(* Logix 5000 project; controller PLC_MCC1300_75F1 vendor 1 type 14 code 166 rev 32.11; software revision 32.04; part 75 of 83 *)
(* tags used below, declared in another part *)
   AUX_tBufferPlate_NULL : UDT_BufferPlate;
   AUX_tHMI_Lite_NULL : UDT_HMI_LITE;
   CONST_rgdDestMask : DINT[32];   // Destination Mask
   CONST_tPlant : UDT_PLANT_CONSTANTS;
   GP_OB_InitializeMain : GP_OB_Initialize;
   GP_PosWindow : GP_PosWindow;
   GP_RampManagement : GP_RampManagement;
   GP_RampSpace : GP_RampSpace;
   M30xTrimDeck : MAC_TrimmingDeck[5];
   M30xTrimDeck_HMR : MAC_TrimmingDeck_HMR[5];
   M30xTrimDeck_HMW : MAC_TrimmingDeck_HMW[5];
   M30xTrimWheel : MAC_TrimmingWheels[5];
   M30xTrimWheel_HMW : MAC_TrimmingWheels_HMW[5];
   M311_Data : UDT_Convoy_SL;
   M311A_Data : UDT_Convoy_SL;
   Sbr_IN_dCapIndex : DINT;
   Sbr_IN_dConveyor : DINT;
   Sbr_IN_DestinationCullet : DINT;
   Sbr_IN_DestinationID : DINT;
   Sbr_IN_dIndexHead : DINT;
   Sbr_IN_dMaskAllowed : DINT;
   Sbr_IN_Position : DINT;
   Sbr_IN_PosStart : DINT;
   Sbr_IN_PosStop : DINT;
   Sbr_IN_ReasonID : DINT;
   Sbr_IN_xHeadPos : BOOL;
   Sbr_IN_xSendAllCullet : BOOL;
   Sbr_INO_DestinationLite : DINT;
   Sbr_INO_tConvoy_SL : UDT_Convoy_SL;
   Sbr_OUT_dIndexTail : DINT;
   Sbr_OUT_ReqRot_CCW : BOOL;
   Sbr_OUT_ReqRot_CW : BOOL;
   TMP_d : DINT;
   TMP_d2 : DINT;
   TMP_dAccSpace : DINT;
   TMP_dActualSpeed : DINT;
   TMP_dBufferSize : DINT;
   TMP_dCap : DINT;
   TMP_dCapNextConvoy : DINT;
   TMP_dConveyorLength : DINT;
   TMP_dConvoySearchMax : DINT;
   TMP_dCountDest : DINT;
   TMP_dCulletMask : DINT;
   TMP_dDecSpace : DINT;
   TMP_dHeadMax : DINT;
   TMP_dHeadPosition_mm : DINT;
   TMP_dIndex : DINT;
   TMP_dIndex2 : DINT;
   TMP_dIndex3 : DINT;
   TMP_dIndex4 : DINT;
   TMP_dIndexCap : DINT;
   TMP_dIndexCapConv : DINT;
   TMP_dIndexConv : DINT;
   TMP_dIndexMotor : DINT;
   TMP_dIndexNext : DINT;
   TMP_dIndexPlate : DINT;
   TMP_dLastConv : DINT;
   TMP_dLastConvTail : DINT;
   TMP_dLineSize : DINT;
   TMP_dLite : DINT;
   TMP_dLiteInv : DINT;
   TMP_dManualTargetPos : DINT;
   TMP_dMask : DINT;
   TMP_dMaxCap : DINT;
   TMP_dMaxLite : DINT;
   TMP_dMinTail : DINT;
   TMP_dNextCap : DINT;
   TMP_dPointerCap : DINT;
   TMP_dPos_cmm : DINT;
   TMP_dPosHead_cmm : DINT;
   TMP_dPosTail_cmm : DINT;
   TMP_dRampMotor : DINT;
   TMP_dStepAdvMotor : DINT;
   TMP_dTotalLength : DINT;
   TMP_dWidth_mm : DINT;
   TMP_IdxLite : DINT;
   TMP_OUT_xPlateEndTracking : BOOL;
   TMP_rgdIndexC : DINT[4];
   TMP_string : STRING;
   TMP_xCenterFound : BOOL;
   TMP_xLastModalityLoadBwd : BOOL;
   TMP_xLastModalityUnloadBwd : BOOL;
   TMP_xMinTailFound : BOOL;
   TMP_xPlateFound : BOOL;
   TMP_xPlateOnConvoyOnNextConveyor : BOOL;
   TMP_xPresenceAlternative : BOOL;
   TMP_xPresenceDestination : BOOL;
   TMP_xPresenceSecondDestination : BOOL;
   TMP_xRun : BOOL;
   TMP_xTailFound : BOOL;
   TMP_xYInversionLite : BOOL;
   TMP_xYWithBarycenter : BOOL;
   xAlwaysOFF : BOOL;
   Z300_BufferPlate : UDT_LINE_BUFFER_PLATE;
   Z300_Conveyor : UDT_StandConv[29];
   Z300_Conveyor_Conf : UDT_Conveyor_Config[29];
   Z300_dEndTrackingPosition : DINT;
   Z300_dStartTrackingPosition : DINT;
   Z300_LineTracking : UDT_LINE_TRACKING;
   Z300_Scada_Continuous : UDT_HMI_LINE_PLATE;
   Z301 : MAC_Zone_ML;
(* MainProgram, continued *)

   12: XIC(M30xTrimDeck_HMR[TMP_dIndex].xControlWidthEnabled)XIC(M30xTrimDeck[TMP_dIndex].ST_xOutputEnable)[XIC(M30xTrimDeck[TMP_dIndex].INPUT_xSATrimDeckToInternal.0) ,XIC(M30xTrimDeck[TMP_dIndex].INPUT_xSATrimDeckToInternal.10) ]ONS(M30xTrimDeck[TMP_dIndex].OSR_xOpSideToInternal)XIO(M30xTrimDeck[TMP_dIndex].INPUT_xSQTrimDeckInternalStop.0)GRT(M30xTrimDeck_HMR[TMP_dIndex].rgdPosition_cmm[0],M30xTrimDeck[TMP_dIndex].CONF_dTrimDeckMinPos_cmm[0])GRT(M30xTrimDeck_HMR[TMP_dIndex].dDistBetweenSides_cmm,M30xTrimDeck[TMP_dIndex].CONF_dTrimDeckMinRange_cmm)SUB(M30xTrimDeck_HMR[TMP_dIndex].rgdOffsetEachSide_cmm[0],M30xTrimDeck_HMW[TMP_dIndex].dOffsetOpSide_cmm,M30xTrimDeck_HMR[TMP_dIndex].rgdOffsetEachSide_cmm[0]);
   13: XIC(M30xTrimDeck_HMR[TMP_dIndex].xControlWidthEnabled)XIC(M30xTrimDeck[TMP_dIndex].ST_xOutputEnable)[XIC(M30xTrimDeck[TMP_dIndex].INPUT_xSATrimDeckToExternal.1) ,XIC(M30xTrimDeck[TMP_dIndex].INPUT_xSATrimDeckToExternal.11) ]ONS(M30xTrimDeck[TMP_dIndex].OSR_xOppOpSideToExternal)XIO(M30xTrimDeck[TMP_dIndex].INPUT_xSQTrimDeckExternalStop.1)LES(M30xTrimDeck_HMR[TMP_dIndex].rgdPosition_cmm[1],M30xTrimDeck[TMP_dIndex].CONF_dTrimDeckMaxPos_cmm[1])LES(M30xTrimDeck_HMR[TMP_dIndex].dDistBetweenSides_cmm,M30xTrimDeck[TMP_dIndex].CONF_dTrimDeckMaxRange_cmm)ADD(M30xTrimDeck_HMR[TMP_dIndex].rgdOffsetEachSide_cmm[1],M30xTrimDeck_HMW[TMP_dIndex].dOffsetOppOpSide_cmm,M30xTrimDeck_HMR[TMP_dIndex].rgdOffsetEachSide_cmm[1]);
   14: XIC(M30xTrimDeck_HMR[TMP_dIndex].xControlWidthEnabled)XIC(M30xTrimDeck[TMP_dIndex].ST_xOutputEnable)[XIC(M30xTrimDeck[TMP_dIndex].INPUT_xSATrimDeckToInternal.1) ,XIC(M30xTrimDeck[TMP_dIndex].INPUT_xSATrimDeckToInternal.11) ]ONS(M30xTrimDeck[TMP_dIndex].OSR_xOppOpSideToInternal)XIO(M30xTrimDeck[TMP_dIndex].INPUT_xSQTrimDeckInternalStop.1)GRT(M30xTrimDeck_HMR[TMP_dIndex].rgdPosition_cmm[1],M30xTrimDeck[TMP_dIndex].CONF_dTrimDeckMinPos_cmm[1])GRT(M30xTrimDeck_HMR[TMP_dIndex].dDistBetweenSides_cmm,M30xTrimDeck[TMP_dIndex].CONF_dTrimDeckMinRange_cmm)SUB(M30xTrimDeck_HMR[TMP_dIndex].rgdOffsetEachSide_cmm[1],M30xTrimDeck_HMW[TMP_dIndex].dOffsetOppOpSide_cmm,M30xTrimDeck_HMR[TMP_dIndex].rgdOffsetEachSide_cmm[1]);
   15: XIC(M30xTrimDeck_HMR[TMP_dIndex].xControlWidthEnabled)XIC(M30xTrimDeck[TMP_dIndex].ST_xOutputEnable)[XIC(M30xTrimDeck[TMP_dIndex].INPUT_xSATrimDeckToOpSide.0) ,XIC(M30xTrimDeck[TMP_dIndex].INPUT_xSATrimDeckToOpSide.1) ]ONS(M30xTrimDeck[TMP_dIndex].OSR_xBothSideToOpSide)XIO(M30xTrimDeck[TMP_dIndex].INPUT_xSQTrimDeckExternalStop.0)LES(M30xTrimDeck_HMR[TMP_dIndex].rgdPosition_cmm[0],M30xTrimDeck[TMP_dIndex].CONF_dTrimDeckMaxPos_cmm[0])XIO(M30xTrimDeck[TMP_dIndex].INPUT_xSQTrimDeckInternalStop.1)GRT(M30xTrimDeck_HMR[TMP_dIndex].rgdPosition_cmm[1],M30xTrimDeck[TMP_dIndex].CONF_dTrimDeckMinPos_cmm[1])SUB(M30xTrimDeck_HMR[TMP_dIndex].dOffsetBothSide_cmm,M30xTrimDeck_HMW[TMP_dIndex].dOffsetOpSide_cmm,M30xTrimDeck_HMR[TMP_dIndex].dOffsetBothSide_cmm);
   16: XIC(M30xTrimDeck_HMR[TMP_dIndex].xControlWidthEnabled)XIC(M30xTrimDeck[TMP_dIndex].ST_xOutputEnable)[XIC(M30xTrimDeck[TMP_dIndex].INPUT_xSATrimDeckToOppOpSide.0) ,XIC(M30xTrimDeck[TMP_dIndex].INPUT_xSATrimDeckToOppOpSide.1) ]ONS(M30xTrimDeck[TMP_dIndex].OSR_xBothSideToOppOpSide)XIO(M30xTrimDeck[TMP_dIndex].INPUT_xSQTrimDeckInternalStop.0)GRT(M30xTrimDeck_HMR[TMP_dIndex].rgdPosition_cmm[0],M30xTrimDeck[TMP_dIndex].CONF_dTrimDeckMinPos_cmm[0])XIO(M30xTrimDeck[TMP_dIndex].INPUT_xSQTrimDeckExternalStop.1)LES(M30xTrimDeck_HMR[TMP_dIndex].rgdPosition_cmm[1],M30xTrimDeck[TMP_dIndex].CONF_dTrimDeckMaxPos_cmm[1])ADD(M30xTrimDeck_HMR[TMP_dIndex].dOffsetBothSide_cmm,M30xTrimDeck_HMW[TMP_dIndex].dOffsetOpSide_cmm,M30xTrimDeck_HMR[TMP_dIndex].dOffsetBothSide_cmm);
   // Request position operator side
   17: [ADD(M30xTrimDeck[TMP_dIndex].AUX_dTarget_cmm[0],M30xTrimDeck_HMR[TMP_dIndex].rgdOffsetEachSide_cmm[0],TMP_d) SUB(TMP_d,M30xTrimDeck_HMR[TMP_dIndex].dOffsetBothSide_cmm,M30xTrimDeck_HMR[TMP_dIndex].rgdTarget_cmm[0]) XIC(xAlwaysOFF) CPT(M30xTrimDeck_HMR[TMP_dIndex].rgdTarget_cmm[0],M30xTrimDeck[TMP_dIndex].AUX_dTarget_cmm[0] + M30xTrimDeck_HMR[TMP_dIndex].rgdOffsetEachSide_cmm[0] - M30xTrimDeck_HMR[TMP_dIndex].dOffsetBothSide_cmm) ,XIC(xAlwaysOFF) XIC(M30xTrimDeck[TMP_dIndex].ST_xJumboInProgress) CPT(M30xTrimDeck_HMR[TMP_dIndex].rgdTarget_cmm[0],M30xTrimDeck_HMR[TMP_dIndex].rgdTarget_cmm[0]) ,XIC(M30xTrimDeck_HMR[TMP_dIndex].xOpeningOnCleaningEnabled) [XIC(Z301.ST_xCleaningAccepted) ,XIC(Z301.OS_xCleaningAccepted) ] MOV(M30xTrimDeck[TMP_dIndex].CONF_dTrimDeckCleanPos_cmm[0],M30xTrimDeck[TMP_dIndex].AUX_dTarget_cmm[0]) MOV(M30xTrimDeck[TMP_dIndex].CONF_dTrimDeckCleanPos_cmm[0],M30xTrimDeck[TMP_dIndex].AUX_dFinalTarget_cmm[0]) MOV(M30xTrimDeck[TMP_dIndex].CONF_dTrimDeckCleanPos_cmm[0],M30xTrimDeck_HMR[TMP_dIndex].rgdTarget_cmm[0]) ,LES(M30xTrimDeck_HMR[TMP_dIndex].rgdTarget_cmm[0],M30xTrimDeck[TMP_dIndex].CONF_dTrimDeckMinPos_cmm[0]) MOV(M30xTrimDeck[TMP_dIndex].CONF_dTrimDeckMinPos_cmm[0],M30xTrimDeck_HMR[TMP_dIndex].rgdTarget_cmm[0]) ,GRT(M30xTrimDeck_HMR[TMP_dIndex].rgdTarget_cmm[0],M30xTrimDeck[TMP_dIndex].CONF_dTrimDeckMaxPos_cmm[0]) MOV(M30xTrimDeck[TMP_dIndex].CONF_dTrimDeckMaxPos_cmm[0],M30xTrimDeck_HMR[TMP_dIndex].rgdTarget_cmm[0]) ,XIC(xAlwaysOFF) GP_PosWindow(GP_PosWindow,M30xTrimDeck_HMR[TMP_dIndex].rgdTarget_cmm[0],M30xTrimDeck_HMR[TMP_dIndex].rgdPosition_cmm[0],M30xTrimDeck[TMP_dIndex].CONF_dTrimDeckDecWindow_cmm[0],0,M30xTrimDeck[TMP_dIndex].ST_xInSlowDownOpSide) ,XIC(xAlwaysOFF) GP_PosWindow(GP_PosWindow,M30xTrimDeck_HMR[TMP_dIndex].rgdTarget_cmm[0],M30xTrimDeck_HMR[TMP_dIndex].rgdPosition_cmm[0],M30xTrimDeck[TMP_dIndex].CONF_dTrimDeckTargetWindow_cmm[0],0,M30xTrimDeck[TMP_dIndex].ST_xInPositionOpSide) ];
   // Request position opposite operator side
   18: [ADD(M30xTrimDeck[TMP_dIndex].AUX_dTarget_cmm[1],M30xTrimDeck_HMR[TMP_dIndex].rgdOffsetEachSide_cmm[1],TMP_d) ADD(TMP_d,M30xTrimDeck_HMR[TMP_dIndex].dOffsetBothSide_cmm,M30xTrimDeck_HMR[TMP_dIndex].rgdTarget_cmm[1]) XIC(xAlwaysOFF) CPT(M30xTrimDeck_HMR[TMP_dIndex].rgdTarget_cmm[1],M30xTrimDeck[TMP_dIndex].AUX_dTarget_cmm[1] + M30xTrimDeck_HMR[TMP_dIndex].rgdOffsetEachSide_cmm[1] + M30xTrimDeck_HMR[TMP_dIndex].dOffsetBothSide_cmm) ,XIC(M30xTrimDeck_HMR[TMP_dIndex].xOpeningOnCleaningEnabled) [XIC(Z301.ST_xCleaningAccepted) ,XIC(Z301.OS_xCleaningAccepted) ] MOV(M30xTrimDeck[TMP_dIndex].CONF_dTrimDeckCleanPos_cmm[0],M30xTrimDeck[TMP_dIndex].AUX_dTarget_cmm[1]) MOV(M30xTrimDeck[TMP_dIndex].CONF_dTrimDeckCleanPos_cmm[0],M30xTrimDeck[TMP_dIndex].AUX_dFinalTarget_cmm[1]) MOV(M30xTrimDeck[TMP_dIndex].CONF_dTrimDeckCleanPos_cmm[1],M30xTrimDeck_HMR[TMP_dIndex].rgdTarget_cmm[1]) ,LES(M30xTrimDeck_HMR[TMP_dIndex].rgdTarget_cmm[1],M30xTrimDeck[TMP_dIndex].CONF_dTrimDeckMinPos_cmm[1]) MOV(M30xTrimDeck[TMP_dIndex].CONF_dTrimDeckMinPos_cmm[1],M30xTrimDeck_HMR[TMP_dIndex].rgdTarget_cmm[1]) ,GRT(M30xTrimDeck_HMR[TMP_dIndex].rgdTarget_cmm[1],M30xTrimDeck[TMP_dIndex].CONF_dTrimDeckMaxPos_cmm[1]) MOV(M30xTrimDeck[TMP_dIndex].CONF_dTrimDeckMaxPos_cmm[1],M30xTrimDeck_HMR[TMP_dIndex].rgdTarget_cmm[1]) ,XIC(xAlwaysOFF) GP_PosWindow(GP_PosWindow,M30xTrimDeck_HMR[TMP_dIndex].rgdTarget_cmm[1],M30xTrimDeck_HMR[TMP_dIndex].rgdPosition_cmm[1],M30xTrimDeck[TMP_dIndex].CONF_dTrimDeckDecWindow_cmm[1],0,M30xTrimDeck[TMP_dIndex].ST_xInSlowDownOppOpSide) ,XIC(xAlwaysOFF) GP_PosWindow(GP_PosWindow,M30xTrimDeck_HMR[TMP_dIndex].rgdTarget_cmm[1],M30xTrimDeck_HMR[TMP_dIndex].rgdPosition_cmm[1],M30xTrimDeck[TMP_dIndex].CONF_dTrimDeckTargetWindow_cmm[1],0,M30xTrimDeck[TMP_dIndex].ST_xInPositionOppOpSide) ];
END_ROUTINE

ROUTINE sbrM311_DecisionRotation   (* structured text *)
   
   //Init
   Sbr_OUT_ReqRot_CW := 0;
   Sbr_OUT_ReqRot_CCW := 0;
   TMP_d := 0;
   TMP_d2 := 0;
   TMP_dMask := CONST_rgdDestMask[0];
   
   //Check qta good lite first cap
   For  TMP_IdxLite := 0 to M311_Data.rgtCap[0].dNumLites -1 by 1 do
   	if M311_Data.rgtCap[0].rgtLite[TMP_IdxLite].tDestination.rgxMain.[TMP_dMask] then
   		TMP_d := TMP_d + 1;
   	end_if;
   end_for;
   
   //Check qta good lite last cap
   if M311A_Data.dTotalCaps > 1 then
   	For  TMP_IdxLite := 0 to M311_Data.rgtCap[0].dNumLites -1 by 1 do
   		if M311_Data.rgtCap[M311A_Data.dTotalCaps - 1].rgtLite[TMP_IdxLite].tDestination.rgxMain.[TMP_dMask] then
   			TMP_d2 := TMP_d2 + 1;
   		end_if;
   	end_for;
   end_if;
   
   //Confront qta
   If TMP_d <= TMP_d2 then
   	Sbr_OUT_ReqRot_CW := 1;
   else
   	Sbr_OUT_ReqRot_CCW := 1;
   end_if;
   
END_ROUTINE

ROUTINE sbrPutLinkConvoy   (* structured text *)
   
   // Reset all indexes
   TMP_dIndex := 0;
   TMP_dIndex2 := 0;
   TMP_dIndex3 := 0;
   TMP_dIndex4 := 0;
   
   TMP_dIndex := TMP_rgdIndexC[0];
   IF TMP_rgdIndexC[1] > 0 THEN
   	TMP_dIndex2 := TMP_rgdIndexC[1];
   END_IF;
   IF TMP_rgdIndexC[2] > 0 THEN
   	TMP_dIndex3 := TMP_rgdIndexC[2];
   END_IF;
   IF TMP_rgdIndexC[3] > 0 THEN
   	TMP_dIndex4 := TMP_rgdIndexC[3];
   END_IF;
   
   // Set convoy index links and length
   Z300_BufferPlate.rgtPlate[TMP_dIndex].tTracking.dPreviousCapIndex := 0;
   Z300_BufferPlate.rgtPlate[TMP_dIndex].tData.rgtCap[0].dConvTotLength_cmm := Z300_BufferPlate.rgtPlate[TMP_dIndex].tData.rgtCap[0].dLength_cmm;
   IF TMP_dIndex2 > 0 THEN
   	Z300_BufferPlate.rgtPlate[TMP_dIndex].tData.dNextCapIndex := TMP_dIndex2;
   	Z300_BufferPlate.rgtPlate[TMP_dIndex].tTracking.dNextCapIndex := TMP_dIndex2;
   	Z300_BufferPlate.rgtPlate[TMP_dIndex2].tTracking.dPreviousCapIndex := TMP_dIndex;
   	Z300_BufferPlate.rgtPlate[TMP_dIndex2].tTracking.dNextCapIndex := 0;
   	Z300_BufferPlate.rgtPlate[TMP_dIndex].tData.rgtCap[0].dConvTotLength_cmm := Z300_BufferPlate.rgtPlate[TMP_dIndex].tData.rgtCap[0].dConvTotLength_cmm + Z300_BufferPlate.rgtPlate[TMP_dIndex].tData.rgtCap[0].dReqGapForConv_cmm + Z300_BufferPlate.rgtPlate[TMP_dIndex2].tData.rgtCap[0].dLength_cmm;
   	Z300_BufferPlate.rgtPlate[TMP_dIndex2].tData.rgtCap[0].dConvTotLength_cmm := Z300_BufferPlate.rgtPlate[TMP_dIndex].tData.rgtCap[0].dConvTotLength_cmm;
   	IF TMP_dIndex3 > 0 THEN
   		Z300_BufferPlate.rgtPlate[TMP_dIndex2].tData.dNextCapIndex := TMP_dIndex3;
   		Z300_BufferPlate.rgtPlate[TMP_dIndex2].tTracking.dNextCapIndex := TMP_dIndex3;
   		Z300_BufferPlate.rgtPlate[TMP_dIndex3].tTracking.dPreviousCapIndex := TMP_dIndex2;
   		Z300_BufferPlate.rgtPlate[TMP_dIndex3].tTracking.dNextCapIndex := 0;
   		Z300_BufferPlate.rgtPlate[TMP_dIndex].tData.rgtCap[0].dConvTotLength_cmm := Z300_BufferPlate.rgtPlate[TMP_dIndex].tData.rgtCap[0].dConvTotLength_cmm + Z300_BufferPlate.rgtPlate[TMP_dIndex2].tData.rgtCap[0].dReqGapForConv_cmm + Z300_BufferPlate.rgtPlate[TMP_dIndex3].tData.rgtCap[0].dLength_cmm;
   		Z300_BufferPlate.rgtPlate[TMP_dIndex2].tData.rgtCap[0].dConvTotLength_cmm := Z300_BufferPlate.rgtPlate[TMP_dIndex].tData.rgtCap[0].dConvTotLength_cmm;
   		Z300_BufferPlate.rgtPlate[TMP_dIndex3].tData.rgtCap[0].dConvTotLength_cmm := Z300_BufferPlate.rgtPlate[TMP_dIndex].tData.rgtCap[0].dConvTotLength_cmm;
   		IF TMP_dIndex4 > 0 THEN
   			Z300_BufferPlate.rgtPlate[TMP_dIndex3].tData.dNextCapIndex := TMP_dIndex4;
   			Z300_BufferPlate.rgtPlate[TMP_dIndex3].tTracking.dNextCapIndex := TMP_dIndex4;
   			Z300_BufferPlate.rgtPlate[TMP_dIndex4].tTracking.dPreviousCapIndex := TMP_dIndex3;
   			Z300_BufferPlate.rgtPlate[TMP_dIndex4].tTracking.dNextCapIndex := 0;
   			Z300_BufferPlate.rgtPlate[TMP_dIndex].tData.rgtCap[0].dConvTotLength_cmm := Z300_BufferPlate.rgtPlate[TMP_dIndex].tData.rgtCap[0].dConvTotLength_cmm + Z300_BufferPlate.rgtPlate[TMP_dIndex3].tData.rgtCap[0].dReqGapForConv_cmm + Z300_BufferPlate.rgtPlate[TMP_dIndex4].tData.rgtCap[0].dLength_cmm;
   			Z300_BufferPlate.rgtPlate[TMP_dIndex2].tData.rgtCap[0].dConvTotLength_cmm := Z300_BufferPlate.rgtPlate[TMP_dIndex].tData.rgtCap[0].dConvTotLength_cmm;
   			Z300_BufferPlate.rgtPlate[TMP_dIndex3].tData.rgtCap[0].dConvTotLength_cmm := Z300_BufferPlate.rgtPlate[TMP_dIndex].tData.rgtCap[0].dConvTotLength_cmm;
   			Z300_BufferPlate.rgtPlate[TMP_dIndex4].tData.rgtCap[0].dConvTotLength_cmm := Z300_BufferPlate.rgtPlate[TMP_dIndex].tData.rgtCap[0].dConvTotLength_cmm;
   		END_IF;
   	END_IF;
   END_IF;
   
END_ROUTINE

ROUTINE sbrRedestConvoyCapZC   (* structured text *)
   
   SBR(Sbr_IN_dCapIndex,Sbr_INO_DestinationLite,Sbr_IN_dMaskAllowed,Sbr_IN_xSendAllCullet,Sbr_IN_DestinationCullet);
   
   
   FOR TMP_dLite := 0 TO Z300_BufferPlate.rgtPlate[Sbr_IN_dCapIndex].tData.rgtCap[0].dNumLites - 1 DO
   	IF Z300_BufferPlate.rgtPlate[Sbr_IN_dCapIndex].tData.rgtCap[0].rgtLite[TMP_dLite].dID <> 0 THEN
   		IF (Z300_BufferPlate.rgtPlate[Sbr_IN_dCapIndex].tData.rgtCap[0].rgtLite[TMP_dLite].tDestination.rgxMain = Sbr_INO_DestinationLite) THEN
   			Z300_BufferPlate.rgtPlate[Sbr_IN_dCapIndex].tData.rgtCap[0].rgtLite[TMP_dLite].tDestination.rgxMain := 0;
   			//filter alternative destinations
   			Z300_BufferPlate.rgtPlate[Sbr_IN_dCapIndex].tData.rgtCap[0].rgtLite[TMP_dLite].tDestination.rgxAlternative := Z300_BufferPlate.rgtPlate[Sbr_IN_dCapIndex].tData.rgtCap[0].rgtLite[TMP_dLite].tDestination.rgxAlternative AND Sbr_IN_dMaskAllowed;
   			IF Sbr_IN_xSendAllCullet OR (Z300_BufferPlate.rgtPlate[Sbr_IN_dCapIndex].tData.rgtCap[0].rgtLite[TMP_dLite].tDestination.rgxAlternative = 0) THEN
   				Z300_BufferPlate.rgtPlate[Sbr_IN_dCapIndex].tData.rgtCap[0].rgtLite[TMP_dLite].tDestination.rgxMain := Sbr_IN_DestinationCullet;
   			ELSE
   				FOR TMP_dIndex := 0 TO 31 DO
   					IF (Z300_BufferPlate.rgtPlate[Sbr_IN_dCapIndex].tData.rgtCap[0].rgtLite[TMP_dLite].tDestination.rgxMain = 0) AND Z300_BufferPlate.rgtPlate[Sbr_IN_dCapIndex].tData.rgtCap[0].rgtLite[TMP_dLite].tDestination.rgxAlternative.[TMP_dIndex] THEN
   						Z300_BufferPlate.rgtPlate[Sbr_IN_dCapIndex].tData.rgtCap[0].rgtLite[TMP_dLite].tDestination.rgxMain.[TMP_dIndex] := 1;
   						Z300_BufferPlate.rgtPlate[Sbr_IN_dCapIndex].tData.rgtCap[0].rgtLite[TMP_dLite].tDestination.rgxAlternative.[TMP_dIndex] := 0;
   					END_IF;
   				END_FOR;
   			END_IF;
   		END_IF;
   	END_IF;
   END_FOR;
   
   IF (Z300_BufferPlate.rgtPlate[Sbr_IN_dCapIndex].tData.dTotalCaps > 1) AND (Z300_BufferPlate.rgtPlate[Sbr_IN_dCapIndex].tTracking.dNextCapIndex > 0) THEN
   	JSR(sbrRedestConvoyCapZC,5,Z300_BufferPlate.rgtPlate[Sbr_IN_dCapIndex].tTracking.dNextCapIndex,Sbr_INO_DestinationLite,Sbr_IN_dMaskAllowed,Sbr_IN_xSendAllCullet,Sbr_IN_DestinationCullet);
   END_IF;
   
END_ROUTINE

ROUTINE sbrRedestConvoySL   (* structured text *)
   
   SBR(Sbr_INO_tConvoy_SL,Sbr_INO_DestinationLite,Sbr_IN_dMaskAllowed,Sbr_IN_xSendAllCullet,Sbr_IN_DestinationCullet);
   
   SIZE(Sbr_INO_tConvoy_SL.rgtCap[0],0,TMP_dMaxCap);
   SIZE(Sbr_INO_tConvoy_SL.rgtCap[0].rgtLite[0],0,TMP_dMaxLite);
   
   FOR TMP_dCap := 0 TO TMP_dMaxCap - 1 DO
   	FOR TMP_dLite := 0 TO TMP_dMaxLite - 1 DO
   		IF Sbr_INO_tConvoy_SL.rgtCap[TMP_dCap].rgtLite[TMP_dLite].dID <> 0 THEN
   			IF Sbr_INO_tConvoy_SL.rgtCap[TMP_dCap].rgtLite[TMP_dLite].tDestination.rgxMain = Sbr_INO_DestinationLite THEN
   				Sbr_INO_tConvoy_SL.rgtCap[TMP_dCap].rgtLite[TMP_dLite].tDestination.rgxMain := 0;
   				//filter alternative destinations
   				Sbr_INO_tConvoy_SL.rgtCap[TMP_dCap].rgtLite[TMP_dLite].tDestination.rgxAlternative := Sbr_INO_tConvoy_SL.rgtCap[TMP_dCap].rgtLite[TMP_dLite].tDestination.rgxAlternative AND Sbr_IN_dMaskAllowed;
   				IF Sbr_IN_xSendAllCullet OR (Sbr_INO_tConvoy_SL.rgtCap[TMP_dCap].rgtLite[TMP_dLite].tDestination.rgxAlternative = 0) THEN
   					Sbr_INO_tConvoy_SL.rgtCap[TMP_dCap].rgtLite[TMP_dLite].tDestination.rgxMain := Sbr_IN_DestinationCullet;
   				ELSE
   					FOR TMP_dIndex := 0 TO 31 DO
   						IF (Sbr_INO_tConvoy_SL.rgtCap[TMP_dCap].rgtLite[TMP_dLite].tDestination.rgxMain = 0) AND Sbr_INO_tConvoy_SL.rgtCap[TMP_dCap].rgtLite[TMP_dLite].tDestination.rgxAlternative.[TMP_dIndex] THEN
   							Sbr_INO_tConvoy_SL.rgtCap[TMP_dCap].rgtLite[TMP_dLite].tDestination.rgxMain.[TMP_dIndex] := 1;
   							Sbr_INO_tConvoy_SL.rgtCap[TMP_dCap].rgtLite[TMP_dLite].tDestination.rgxAlternative.[TMP_dIndex] := 0;
   						END_IF;
   					END_FOR;
   				END_IF;
   			END_IF;
   		END_IF;
   	END_FOR;
   END_FOR;
   
   RET(Sbr_INO_tConvoy_SL);
   
END_ROUTINE

ROUTINE sbrResetLinkConvoy   (* structured text *)
   
   FOR TMP_dIndex := 0 TO 3 DO
   	TMP_rgdIndexC[TMP_dIndex] := 0;
   END_FOR;
   
END_ROUTINE

ROUTINE sbrTrackingConvPresence   (* structured text *)
   
   FOR TMP_dIndexConv := 0 TO CONST_tPlant.dNumOfConveyors - 1 DO
       IF Z300_LineTracking.rgtTrkConv[TMP_dIndexConv].dIndexCaps <> 0  THEN //Plate on Conveyor
           TMP_dHeadMax := 0;
           TMP_dMinTail := Z300_LineTracking.rgtTrkConv[TMP_dIndexConv].dEndPosition_cmm;
           TMP_xMinTailFound := 0;
           FOR TMP_dCap := 0 TO Z300_LineTracking.rgtTrkConv[TMP_dIndexConv].dIndexCaps - 1 DO
               //Take Pointer
               TMP_dPointerCap := Z300_LineTracking.rgtTrkConv[TMP_dIndexConv].Cap[TMP_dCap].dPointer;
               //Check Plate id Convoy Presence on next Conveyor
               TMP_xPlateOnConvoyOnNextConveyor := 0;
               //Convoy Presence Check for the next conveyor
               IF Z300_BufferPlate.rgtPlate[TMP_dPointerCap].tTracking.dPreviousCapIndex <> 0 AND TMP_dIndexConv + TMP_dIndexNext < CONST_tPlant.dNumOfConveyors THEN
                   TMP_dConvoySearchMax := 1;
                   TMP_dTotalLength := 0;
                   //Search if the length is more that the Next (search up to three conveyors next)
                   FOR TMP_dIndexNext := 1 TO 3 DO
                       IF TMP_dIndexConv + TMP_dIndexNext < CONST_tPlant.dNumOfConveyors THEN
                           IF Z300_BufferPlate.rgtPlate[TMP_dPointerCap].tData.dGapCaps_cmm >= Z300_LineTracking.rgtTrkConv[TMP_dIndexConv + TMP_dIndexNext].dLengthConveyor + TMP_dTotalLength THEN
                               TMP_dConvoySearchMax := TMP_dIndexNext + 1;
                           ELSE
                               EXIT;
                           END_IF;
                           TMP_dTotalLength := Z300_LineTracking.rgtTrkConv[TMP_dIndexConv + TMP_dIndexNext].dLengthConveyor;
                       END_IF;
                   END_FOR;
   
                   FOR TMP_dIndexNext := 1 TO TMP_dConvoySearchMax DO
                       IF TMP_dIndexConv + TMP_dIndexNext < CONST_tPlant.dNumOfConveyors THEN
                           IF Z300_LineTracking.rgtTrkConv[TMP_dIndexConv + TMP_dIndexNext].dIndexCaps <> 0 THEN //Enter to Search in case of  Glass
                               FOR TMP_dCapNextConvoy := 0 TO Z300_LineTracking.rgtTrkConv[TMP_dIndexConv].dIndexCaps DO //Cehck if there are the same Index Plate
   								IF (TMP_dCapNextConvoy < CONST_tPlant.dNumCapsConveyor) THEN
   	                                TMP_xPlateOnConvoyOnNextConveyor := 0;
   									IF Z300_BufferPlate.rgtPlate[TMP_dPointerCap].tTracking.dPreviousCapIndex = Z300_LineTracking.rgtTrkConv[TMP_dIndexConv + TMP_dIndexNext].Cap[TMP_dCapNextConvoy].dPointer THEN
   										TMP_xPlateOnConvoyOnNextConveyor := 1;
   									END_IF;
   	                                IF TMP_dIndexNext <> 1 THEN
   	                                    Z300_LineTracking.rgtTrkConv[TMP_dIndexConv + TMP_dIndexNext - 1].xPlateConvPreviousNext := TMP_xPlateOnConvoyOnNextConveyor;
   	                                END_IF;
   	                                IF TMP_xPlateOnConvoyOnNextConveyor OR (Z300_LineTracking.rgtTrkConv[TMP_dIndexConv + TMP_dIndexNext].Cap[TMP_dCapNextConvoy].dPointer = 0) THEN
   	                                    EXIT; //EXit When Found the Value or if the index is 0
   	                                END_IF;
   								END_IF;
                               END_FOR;
                           END_IF;
                       END_IF;
                   END_FOR;
               END_IF;
   
               //Check The Max and The minimun Head and Tail
   			////IF TMP_dHeadMax <= Z300_LineTracking.rgtTrkConv[TMP_dIndexConv].Cap[TMP_dCap].dHeadPos_cmm AND NOT TMP_xPlateOnConvoyOnNextConveyor THEN
               IF TMP_dHeadMax <= Z300_LineTracking.rgtTrkConv[TMP_dIndexConv].Cap[TMP_dCap].dHeadPos_cmm AND (NOT TMP_xPlateOnConvoyOnNextConveyor) AND (NOT Z300_BufferPlate.rgtPlate[TMP_dPointerCap].tTracking.xNotConsConvTrk) THEN
                   TMP_dHeadMax := Z300_LineTracking.rgtTrkConv[TMP_dIndexConv].Cap[TMP_dCap].dHeadPos_cmm;
               END_IF;
               TMP_dPointerCap := Z300_LineTracking.rgtTrkConv[TMP_dIndexConv].Cap[TMP_dCap].dPointer;
               IF  TMP_dMinTail >= Z300_LineTracking.rgtTrkConv[TMP_dIndexConv].Cap[TMP_dCap].dTailPos_cmm AND Z300_LineTracking.rgtTrkConv[TMP_dIndexConv].Cap[TMP_dCap].xTail
                   AND (Z300_BufferPlate.rgtPlate[TMP_dPointerCap].tTracking.dNextCapIndex = 0) THEN
                   TMP_dMinTail := Z300_LineTracking.rgtTrkConv[TMP_dIndexConv].Cap[TMP_dCap].dTailPos_cmm;
                   TMP_xMinTailFound := 1;
               END_IF;
   
   			//Double motor management
   			IF Z300_Conveyor_Conf[TMP_dIndexConv].dMotorNumber > 0 THEN
                   TMP_dRampMotor := Z300_BufferPlate.rgtPlate[TMP_dPointerCap].tTracking.dIndexMotorStepAdv;
               ELSE //One motor presence considerate the plate on the first
                       TMP_dRampMotor := 0;
               END_IF;
   
               //Plate passage Downstream
               Z300_LineTracking.rgtTrkConv[TMP_dIndexConv].xPlatePassageNext := Z300_LineTracking.rgtTrkConv[TMP_dIndexConv].xPlatePassageNext OR
               ((Z300_LineTracking.rgtTrkConv[TMP_dIndexConv].Cap[TMP_dCap].dHeadPosConv_cmm
   			+ Z300_LineTracking.rgtTrkConv[TMP_dIndexConv].dActualRamp_cmm[0] > Z300_LineTracking.rgtTrkConv[TMP_dIndexConv].dLengthConveyor
               OR (Z300_LineTracking.rgtTrkConv[TMP_dIndexConv].Cap[TMP_dCap].xPresence AND NOT(Z300_LineTracking.rgtTrkConv[TMP_dIndexConv].Cap[TMP_dCap].xHead))
               OR TMP_xPlateOnConvoyOnNextConveyor  OR Z300_LineTracking.rgtTrkConv[TMP_dIndexConv].xPlatePassageNext
   			OR Z300_LineTracking.rgtTrkConv[TMP_dIndexConv].xPlateConvPreviousNext)
               AND ((NOT Z300_BufferPlate.rgtPlate[TMP_dPointerCap].tTracking.xNotConsConvTrk) OR TMP_dIndexConv < Z300_BufferPlate.rgtPlate[TMP_dPointerCap].tTracking.dIndexConvNotCons));
   
               IF TMP_dIndexConv + 1 < CONST_tPlant.dNumOfConveyors THEN
                   Z300_LineTracking.rgtTrkConv[TMP_dIndexConv + 1].xPlatePassagePrevious := Z300_LineTracking.rgtTrkConv[TMP_dIndexConv].xPlatePassageNext;
               END_IF;
               //Glass Presence
               Z300_LineTracking.rgtTrkConv[TMP_dIndexConv].xGlassPresence := Z300_LineTracking.rgtTrkConv[TMP_dIndexConv].xGlassPresence OR
   			(Z300_LineTracking.rgtTrkConv[TMP_dIndexConv].Cap[TMP_dCap].xPresence AND ((NOT Z300_BufferPlate.rgtPlate[TMP_dPointerCap].tTracking.xNotConsConvTrk)
               OR TMP_dIndexConv < Z300_BufferPlate.rgtPlate[TMP_dPointerCap].tTracking.dIndexConvNotCons));
   
           END_FOR;
           Z300_LineTracking.rgtTrkConv[TMP_dIndexConv].dHeadPosition_cmm:= TMP_dHeadMax;
           IF TMP_xMinTailFound THEN
               Z300_LineTracking.rgtTrkConv[TMP_dIndexConv].dTailPosition_cmm := TMP_dMinTail;
           ELSE
               TMP_dMinTail := 0;
           END_IF;
       ELSIF Z300_LineTracking.rgtTrkConv[TMP_dIndexConv].xPlateConvPreviousNext THEN
           Z300_LineTracking.rgtTrkConv[TMP_dIndexConv].xPlatePassageNext := 1;
           IF TMP_dIndexConv + 1 < CONST_tPlant.dNumOfConveyors THEN
               Z300_LineTracking.rgtTrkConv[TMP_dIndexConv + 1].xPlatePassagePrevious := 1;
           END_IF;
       END_IF;
       Z300_LineTracking.rgtTrkConv[TMP_dIndexConv].xGlassPresCom := Z300_LineTracking.rgtTrkConv[TMP_dIndexConv].xPlatePassagePrevious
   																		OR Z300_LineTracking.rgtTrkConv[TMP_dIndexConv].xGlassPresence;
   	Z300_LineTracking.rgtTrkConv[TMP_dIndexConv].xHeadPresenceConv := Z300_LineTracking.rgtTrkConv[TMP_dIndexConv].dHeadPosition_cmm <> 0;
   END_FOR;
   
END_ROUTINE

ROUTINE sbrTrackingConvStep   (* ladder *)
   // #####_COSTANTS_#####
   0: MOV(0,TMP_dIndexMotor);
   // #####_LOOP FOR MOTOR_#####
   1: LBL(AuxLoop)NOP();
   2: XIC(Z300_Conveyor[TMP_dIndexConv].ST_xConveyorOutRun)XIC(Z300_Conveyor[TMP_dIndexConv].ST_rgxOutMotorRunSgm.[TMP_dIndexMotor])XIO(Z300_Conveyor[TMP_dIndexConv].ST_xDriveInDec)XIC(Z300_Conveyor[TMP_dIndexConv].ST_xAxleReadyToMoveDelayed)OTE(TMP_xRun);
   3: GP_RampManagement(GP_RampManagement,TMP_xRun,Z300_Conveyor[TMP_dIndexConv].AUX_rgdCurrentSpeed_mm_min[TMP_dIndexMotor],Z300_Conveyor[TMP_dIndexConv].AUX_rgrAcc_m_s2[TMP_dIndexMotor],Z300_Conveyor[TMP_dIndexConv].AUX_rgrDec_m_s2[TMP_dIndexMotor],GP_OB_InitializeMain.OUT_dExecutionTime_ms,Z300_Conveyor[TMP_dIndexConv].AUX_rgrSpeedIncrement_mm_min[TMP_dIndexMotor],Z300_Conveyor[TMP_dIndexConv].AUX_rgdStepAdvancement_cmm[TMP_dIndexMotor],Z300_Conveyor[TMP_dIndexConv].ST_rgxRampInProgress.[TMP_dIndexMotor],Z300_Conveyor[TMP_dIndexConv].ST_rgxAccInProgress.[TMP_dIndexMotor],Z300_Conveyor[TMP_dIndexConv].ST_rgxDecInProgress.[TMP_dIndexMotor],Z300_Conveyor[TMP_dIndexConv].AUX_rgrReminderStep[TMP_dIndexMotor]);
   4: MOV(Z300_Conveyor[TMP_dIndexConv].AUX_rgdCurrentSpeed_mm_min[TMP_dIndexMotor],TMP_dActualSpeed);
   5: XIO(Z300_Conveyor[TMP_dIndexConv].ST_xRotationFeedback)XIO(Z300_Conveyor[TMP_dIndexConv].ST_rgxDecInProgress.[TMP_dIndexMotor])MOV(0,TMP_dActualSpeed);
   6: GP_RampSpace(GP_RampSpace,Z300_Conveyor[TMP_dIndexConv].AUX_rgrAcc_m_s2[TMP_dIndexMotor],Z300_Conveyor[TMP_dIndexConv].AUX_rgrDec_m_s2[TMP_dIndexMotor],TMP_dActualSpeed,TMP_dAccSpace,TMP_dDecSpace);
   7: MOV(Z300_Conveyor[TMP_dIndexConv].AUX_rgdStepAdvancement_cmm[TMP_dIndexMotor],Z300_LineTracking.rgtTrkConv[TMP_dIndexConv].dStepAdv_cmm[TMP_dIndexMotor]);
   8: MOV(TMP_dDecSpace,Z300_LineTracking.rgtTrkConv[TMP_dIndexConv].dActualRamp_cmm[TMP_dIndexMotor]);
   9: MOV(Z300_Conveyor_Conf[TMP_dIndexConv].dLengthConveyor_cmm,Z300_LineTracking.rgtTrkConv[TMP_dIndexConv].dLengthConveyor);
   10: LES(TMP_dIndexMotor,Z300_Conveyor_Conf[TMP_dIndex].dMotorNumber)ADD(TMP_dIndexMotor,1,TMP_dIndexMotor)JMP(AuxLoop);
END_ROUTINE

ROUTINE sbrTrackingDeleteConvoy   (* structured text *)
   
   SBR(Sbr_IN_dCapIndex);
   
   TMP_dNextCap := 0;
   IF Z300_BufferPlate.rgtPlate[Sbr_IN_dCapIndex].tData.dTotalCaps > 1 THEN
   	TMP_dNextCap := Z300_BufferPlate.rgtPlate[Sbr_IN_dCapIndex].tTracking.dNextCapIndex;
   END_IF;
   
   // Delete this cap
   COP(AUX_tBufferPlate_NULL,Z300_BufferPlate.rgtPlate[Sbr_IN_dCapIndex],1);
   IF TMP_dNextCap > 0 THEN
   	// Call recursively to next cap
   	JSR(sbrTrackingDeleteConvoy,1,TMP_dNextCap);
   END_IF;
   
END_ROUTINE

ROUTINE sbrTrackingHideConvPresence   (* structured text *)
   
   SBR(Sbr_IN_dCapIndex,Sbr_IN_dConveyor);
   
   Z300_BufferPlate.rgtPlate[Sbr_IN_dCapIndex].tTracking.xNotConsConvTrk := 1;
   IF Z300_BufferPlate.rgtPlate[Sbr_IN_dCapIndex].tTracking.dIndexConvNotCons > Sbr_IN_dConveyor THEN
   	Z300_BufferPlate.rgtPlate[Sbr_IN_dCapIndex].tTracking.dIndexConvNotCons := Sbr_IN_dConveyor;
   END_IF;
   IF (Z300_BufferPlate.rgtPlate[Sbr_IN_dCapIndex].tData.dTotalCaps > 1) AND (Z300_BufferPlate.rgtPlate[Sbr_IN_dCapIndex].tTracking.dNextCapIndex > 0) THEN
   	JSR(sbrTrackingHideConvPresence,2,Z300_BufferPlate.rgtPlate[Sbr_IN_dCapIndex].tTracking.dNextCapIndex,Sbr_IN_dConveyor);
   END_IF;
   
END_ROUTINE

ROUTINE sbrTrackingIndexNotInConvoy   (* ladder *)
   0: XIC(Z300_BufferPlate.rgtPlate[TMP_dIndex].tTracking.xNotConsConvTrk)LEQ(Z300_BufferPlate.rgtPlate[TMP_dIndex].tTracking.dIndexConvNotCons,0)MOV(Z300_BufferPlate.rgtPlate[TMP_dIndex].tTracking.dIndexConvHead,Z300_BufferPlate.rgtPlate[TMP_dIndex].tTracking.dIndexConvNotCons);
   1: XIO(Z300_BufferPlate.rgtPlate[TMP_dIndex].tTracking.xNotConsConvTrk)MOV(0,Z300_BufferPlate.rgtPlate[TMP_dIndex].tTracking.dIndexConvNotCons);
END_ROUTINE

ROUTINE sbrTrackingIndexTailConvoy   (* structured text *)
   
   //Finds tail of convoy in recursive mode
   //Input
   SBR(Sbr_IN_dIndexHead);
   IF Z300_BufferPlate.rgtPlate[Sbr_IN_dIndexHead].tTracking.dNextCapIndex > 0 THEN
   	JSR(sbrTrackingIndexTailConvoy,1,Z300_BufferPlate.rgtPlate[Sbr_IN_dIndexHead].tTracking.dNextCapIndex,Sbr_OUT_dIndexTail);
   ELSE
       Sbr_OUT_dIndexTail := Sbr_IN_dIndexHead;
   END_IF;
   
   //Write output
   RET(Sbr_OUT_dIndexTail);
   
END_ROUTINE

ROUTINE sbrTrackingPlateCleaning   (* structured text *)
   
   SBR(Sbr_IN_PosStart,Sbr_IN_PosStop,Sbr_IN_DestinationID,Sbr_IN_ReasonID);
   COP(TMP_string,TMP_string,1);
   SIZE(Z300_BufferPlate.rgtPlate[0],0,TMP_dBufferSize);
   FOR TMP_dIndex := 1 TO TMP_dBufferSize - 1 DO
   	IF Z300_BufferPlate.rgtPlate[TMP_dIndex].tTracking.dPositionHead_cmm >= Sbr_IN_PosStart
   		AND Z300_BufferPlate.rgtPlate[TMP_dIndex].tTracking.dPositionHead_cmm <= Sbr_IN_PosStop
   			AND Z300_BufferPlate.rgtPlate[TMP_dIndex].tData.dLength_cmm <> 0 THEN
   
   		FOR TMP_dLite := 0 TO Z300_BufferPlate.rgtPlate[0].tData.rgtCap[0].dNumLites - 1 DO
   			IF Z300_BufferPlate.rgtPlate[TMP_dIndex].tData.rgtCap[0].rgtLite[TMP_dLite].dID <> 0 THEN
   				IF Z300_BufferPlate.rgtPlate[TMP_dIndex].tData.rgtCap[0].rgtLite[TMP_dLite].dCulletCause = 0 THEN
   					// Plate redestination message
   					//RP_AddMessageV2(RP_AddMessage,
   					//			0,
   					//			RP_tMessagesCode.Message[8],
   					//			Sbr_IN_DestinationID,
   					//			Z300_BufferPlate.rgtPlate[TMP_dIndex].tData.rgtCap[0].rgtLite[TMP_dLite].dID,
   					//			Z300_BufferPlate.rgtPlate[TMP_dIndex].tData.rgtCap[0].rgtLite[TMP_dLite].dProductionID,
   					//			Sbr_IN_ReasonID,
   					//			0,
   					//			0,
   					//			0,
   					//			0,
   					//			0,
   					//			0,
   					//			RP_tAddMessageBuffer,
   					//			RP_xAddMessageError,
   					//			TMP_string);
   				END_IF;
   				// Plate broken message
   				//RP_AddMessageV2(RP_AddMessage,
   				//				0,
   				//				RP_tMessagesCode.Message[2],
   				//				Sbr_IN_DestinationID,
   				//				Z300_BufferPlate.rgtPlate[TMP_dIndex].tData.rgtCap[0].rgtLite[TMP_dLite].dID,
   				//				Z300_BufferPlate.rgtPlate[TMP_dIndex].tData.rgtCap[0].rgtLite[TMP_dLite].dProductionID,
   				//				0,
   				//				0,
   				//				0,
   				//				0,
   				//				0,
   				//				0,
   				//				0,
   				//				RP_tAddMessageBuffer,
   				//				RP_xAddMessageError,
   				//				TMP_string);
   			END_IF;
   		END_FOR;
   		COP(AUX_tBufferPlate_NULL, Z300_BufferPlate.rgtPlate[TMP_dIndex], 1);
   	END_IF;
   END_FOR;
   
END_ROUTINE

ROUTINE sbrTrackingPositioningDone   (* structured text *)
   
   SBR(Sbr_IN_dCapIndex,Sbr_IN_xHeadPos,Sbr_IN_Position);